screen "752_Profinet_IO_System" 1280x800, template "Top_Header"
   on GenerateScreen: SetTag("UserDiag_HmiData_actIOSystem", 1)
   on ClearScreen: SetTag("UserDiag_HmiData_actIOSystem", -2)
   TextField "Text field_1" at 7,121 size 149x32; Text 'IO Systeme / IO Systems'
   Button "Schaltfläche_64" at 950,700 size 250x80; TextOn 'Reset Übersicht / Reset overview'; TextOff 'Reset Übersicht / Reset overview'
      on Press: function_b14e0dd5("UserDiag_HmiData_ackStates", 0)
   ScreenModuleView "typeDevice_1" at 110,154 size 110x110; ScreenModuleType ""
      on Guid_{11997190-132388}: SetTag("UserDiag_HmiData_actDeviceOfScreen", 1); function_efd93a16("Pop-up_OverviewModules", 0, 0, -1, -1, 2); SetBit("UserDiag_HmiData_ioSlotDiagnosticsLoaded")
      Guid_{11997190-132400} <- "[0]"
      Guid_{11997190-132580} <- "[0]"
   ScreenModuleView "typeDevice_2" at 250,154 size 110x110; ScreenModuleType ""
      on Guid_{11997190-132388}: SetTag("UserDiag_HmiData_actDeviceOfScreen", 2); function_efd93a16("Pop-up_OverviewModules", 0, 0, -1, -1, 2); SetBit("UserDiag_HmiData_ioSlotDiagnosticsLoaded")
      Guid_{11997190-132400} <- "[1]"
      Guid_{11997190-132580} <- "[1]"
   ScreenModuleView "typeDevice_3" at 390,154 size 110x110; ScreenModuleType ""
      on Guid_{11997190-132388}: SetTag("UserDiag_HmiData_actDeviceOfScreen", 3); function_efd93a16("Pop-up_OverviewModules", 0, 0, -1, -1, 2); SetBit("UserDiag_HmiData_ioSlotDiagnosticsLoaded")
      Guid_{11997190-132400} <- "[2]"
      Guid_{11997190-132580} <- "[2]"
   ScreenModuleView "typeDevice_4" at 530,154 size 110x110; ScreenModuleType ""
      on Guid_{11997190-132388}: SetTag("UserDiag_HmiData_actDeviceOfScreen", 4); function_efd93a16("Pop-up_OverviewModules", 0, 0, -1, -1, 2); SetBit("UserDiag_HmiData_ioSlotDiagnosticsLoaded")
      Guid_{11997190-132400} <- "[3]"
      Guid_{11997190-132580} <- "[3]"
   ScreenModuleView "typeDevice_5" at 670,154 size 110x110; ScreenModuleType ""
      on Guid_{11997190-132388}: SetTag("UserDiag_HmiData_actDeviceOfScreen", 5); function_efd93a16("Pop-up_OverviewModules", 0, 0, -1, -1, 2); SetBit("UserDiag_HmiData_ioSlotDiagnosticsLoaded")
      Guid_{11997190-132400} <- "[4]"
      Guid_{11997190-132580} <- "[4]"
   ScreenModuleView "typeDevice_6" at 810,154 size 110x110; ScreenModuleType ""
      on Guid_{11997190-132388}: SetTag("UserDiag_HmiData_actDeviceOfScreen", 6); function_efd93a16("Pop-up_OverviewModules", 0, 0, -1, -1, 2); SetBit("UserDiag_HmiData_ioSlotDiagnosticsLoaded")
      Guid_{11997190-132400} <- "[5]"
      Guid_{11997190-132580} <- "[5]"
   ScreenModuleView "typeDevice_7" at 950,154 size 110x110; ScreenModuleType ""
      on Guid_{11997190-132388}: SetTag("UserDiag_HmiData_actDeviceOfScreen", 7); function_efd93a16("Pop-up_OverviewModules", 0, 0, -1, -1, 2); SetBit("UserDiag_HmiData_ioSlotDiagnosticsLoaded")
      Guid_{11997190-132400} <- "[6]"
      Guid_{11997190-132580} <- "[6]"
   ScreenModuleView "typeDevice_8" at 1090,154 size 110x110; ScreenModuleType ""
      on Guid_{11997190-132388}: SetTag("UserDiag_HmiData_actDeviceOfScreen", 8); function_efd93a16("Pop-up_OverviewModules", 0, 0, -1, -1, 2); SetBit("UserDiag_HmiData_ioSlotDiagnosticsLoaded")
      Guid_{11997190-132400} <- "[7]"
      Guid_{11997190-132580} <- "[7]"
   ScreenModuleView "typeDevice_9" at 110,294 size 110x110; ScreenModuleType ""
      on Guid_{11997190-132388}: SetTag("UserDiag_HmiData_actDeviceOfScreen", 9); function_efd93a16("Pop-up_OverviewModules", 0, 0, -1, -1, 2); SetBit("UserDiag_HmiData_ioSlotDiagnosticsLoaded")
      Guid_{11997190-132400} <- "[8]"
      Guid_{11997190-132580} <- "[8]"
   ScreenModuleView "typeDevice_10" at 250,294 size 110x110; ScreenModuleType ""
      on Guid_{11997190-132388}: SetTag("UserDiag_HmiData_actDeviceOfScreen", 10); function_efd93a16("Pop-up_OverviewModules", 0, 0, -1, -1, 2); SetBit("UserDiag_HmiData_ioSlotDiagnosticsLoaded")
      Guid_{11997190-132400} <- "[9]"
      Guid_{11997190-132580} <- "[9]"
   ScreenModuleView "typeDevice_11" at 390,294 size 110x110; ScreenModuleType ""
      on Guid_{11997190-132388}: SetTag("UserDiag_HmiData_actDeviceOfScreen", 11); function_efd93a16("Pop-up_OverviewModules", 0, 0, -1, -1, 2); SetBit("UserDiag_HmiData_ioSlotDiagnosticsLoaded")
      Guid_{11997190-132400} <- "[10]"
      Guid_{11997190-132580} <- "[10]"
   ScreenModuleView "typeDevice_12" at 530,294 size 110x110; ScreenModuleType ""
      on Guid_{11997190-132388}: SetTag("UserDiag_HmiData_actDeviceOfScreen", 12); function_efd93a16("Pop-up_OverviewModules", 0, 0, -1, -1, 2); SetBit("UserDiag_HmiData_ioSlotDiagnosticsLoaded")
      Guid_{11997190-132400} <- "[11]"
      Guid_{11997190-132580} <- "[11]"
   ScreenModuleView "typeDevice_13" at 670,294 size 110x110; ScreenModuleType ""
      on Guid_{11997190-132388}: SetTag("UserDiag_HmiData_actDeviceOfScreen", 13); function_efd93a16("Pop-up_OverviewModules", 0, 0, -1, -1, 2); SetBit("UserDiag_HmiData_ioSlotDiagnosticsLoaded")
      Guid_{11997190-132400} <- "[12]"
      Guid_{11997190-132580} <- "[12]"
   ScreenModuleView "typeDevice_14" at 810,294 size 110x110; ScreenModuleType ""
      on Guid_{11997190-132388}: SetTag("UserDiag_HmiData_actDeviceOfScreen", 14); function_efd93a16("Pop-up_OverviewModules", 0, 0, -1, -1, 2); SetBit("UserDiag_HmiData_ioSlotDiagnosticsLoaded")
      Guid_{11997190-132400} <- "[13]"
      Guid_{11997190-132580} <- "[13]"
   ScreenModuleView "typeDevice_15" at 950,292 size 110x110; ScreenModuleType ""
      on Guid_{11997190-132388}: SetTag("UserDiag_HmiData_actDeviceOfScreen", 15); function_efd93a16("Pop-up_OverviewModules", 0, 0, -1, -1, 2); SetBit("UserDiag_HmiData_ioSlotDiagnosticsLoaded")
      Guid_{11997190-132400} <- "[14]"
      Guid_{11997190-132580} <- "[14]"
   ScreenModuleView "typeDevice_16" at 1090,294 size 110x110; ScreenModuleType ""
      on Guid_{11997190-132388}: SetTag("UserDiag_HmiData_actDeviceOfScreen", 16); function_efd93a16("Pop-up_OverviewModules", 0, 0, -1, -1, 2); SetBit("UserDiag_HmiData_ioSlotDiagnosticsLoaded")
      Guid_{11997190-132400} <- "[15]"
      Guid_{11997190-132580} <- "[15]"
   ScreenModuleView "typeDevice_17" at 110,434 size 110x110; ScreenModuleType ""
      on Guid_{11997190-132388}: SetTag("UserDiag_HmiData_actDeviceOfScreen", 17); function_efd93a16("Pop-up_OverviewModules", 0, 0, -1, -1, 2); SetBit("UserDiag_HmiData_ioSlotDiagnosticsLoaded")
      Guid_{11997190-132400} <- "[16]"
      Guid_{11997190-132580} <- "[16]"
   ScreenModuleView "typeDevice_18" at 250,434 size 110x110; ScreenModuleType ""
      on Guid_{11997190-132388}: SetTag("UserDiag_HmiData_actDeviceOfScreen", 18); function_efd93a16("Pop-up_OverviewModules", 0, 0, -1, -1, 2); SetBit("UserDiag_HmiData_ioSlotDiagnosticsLoaded")
      Guid_{11997190-132400} <- "[17]"
      Guid_{11997190-132580} <- "[17]"
   ScreenModuleView "typeDevice_19" at 390,434 size 110x110; ScreenModuleType ""
      on Guid_{11997190-132388}: SetTag("UserDiag_HmiData_actDeviceOfScreen", 19); function_efd93a16("Pop-up_OverviewModules", 0, 0, -1, -1, 2); SetBit("UserDiag_HmiData_ioSlotDiagnosticsLoaded")
      Guid_{11997190-132400} <- "[18]"
      Guid_{11997190-132580} <- "[18]"
   ScreenModuleView "typeDevice_20" at 530,434 size 110x110; ScreenModuleType ""
      on Guid_{11997190-132388}: SetTag("UserDiag_HmiData_actDeviceOfScreen", 20); function_efd93a16("Pop-up_OverviewModules", 0, 0, -1, -1, 2); SetBit("UserDiag_HmiData_ioSlotDiagnosticsLoaded")
      Guid_{11997190-132400} <- "[19]"
      Guid_{11997190-132580} <- "[19]"
   ScreenModuleView "typeDevice_21" at 670,434 size 110x110; ScreenModuleType ""
      on Guid_{11997190-132388}: SetTag("UserDiag_HmiData_actDeviceOfScreen", 21); function_efd93a16("Pop-up_OverviewModules", 0, 0, -1, -1, 2); SetBit("UserDiag_HmiData_ioSlotDiagnosticsLoaded")
      Guid_{11997190-132400} <- "[20]"
      Guid_{11997190-132580} <- "[20]"
   ScreenModuleView "typeDevice_22" at 810,434 size 110x110; ScreenModuleType ""
      on Guid_{11997190-132388}: SetTag("UserDiag_HmiData_actDeviceOfScreen", 22); function_efd93a16("Pop-up_OverviewModules", 0, 0, -1, -1, 2); SetBit("UserDiag_HmiData_ioSlotDiagnosticsLoaded")
      Guid_{11997190-132400} <- "[21]"
      Guid_{11997190-132580} <- "[21]"
   ScreenModuleView "typeDevice_23" at 950,434 size 110x110; ScreenModuleType ""
      on Guid_{11997190-132388}: SetTag("UserDiag_HmiData_actDeviceOfScreen", 23); function_efd93a16("Pop-up_OverviewModules", 0, 0, -1, -1, 2); SetBit("UserDiag_HmiData_ioSlotDiagnosticsLoaded")
      Guid_{11997190-132400} <- "[22]"
      Guid_{11997190-132580} <- "[22]"
   ScreenModuleView "typeDevice_24" at 1090,434 size 110x110; ScreenModuleType ""
      on Guid_{11997190-132388}: SetTag("UserDiag_HmiData_actDeviceOfScreen", 24); function_efd93a16("Pop-up_OverviewModules", 0, 0, -1, -1, 2); SetBit("UserDiag_HmiData_ioSlotDiagnosticsLoaded")
      Guid_{11997190-132400} <- "[23]"
      Guid_{11997190-132580} <- "[23]"
   ScreenModuleView "typeDevice_25" at 110,574 size 110x110; ScreenModuleType ""
      on Guid_{11997190-132388}: SetTag("UserDiag_HmiData_actDeviceOfScreen", 25); function_efd93a16("Pop-up_OverviewModules", 0, 0, -1, -1, 2); SetBit("UserDiag_HmiData_ioSlotDiagnosticsLoaded")
      Guid_{11997190-132400} <- "[24]"
      Guid_{11997190-132580} <- "[24]"
   ScreenModuleView "typeDevice_26" at 250,574 size 110x110; ScreenModuleType ""
      on Guid_{11997190-132388}: SetTag("UserDiag_HmiData_actDeviceOfScreen", 26); function_efd93a16("Pop-up_OverviewModules", 0, 0, -1, -1, 2); SetBit("UserDiag_HmiData_ioSlotDiagnosticsLoaded")
      Guid_{11997190-132400} <- "[25]"
      Guid_{11997190-132580} <- "[25]"
   ScreenModuleView "typeDevice_27" at 390,574 size 110x110; ScreenModuleType ""
      on Guid_{11997190-132388}: SetTag("UserDiag_HmiData_actDeviceOfScreen", 27); function_efd93a16("Pop-up_OverviewModules", 0, 0, -1, -1, 2); SetBit("UserDiag_HmiData_ioSlotDiagnosticsLoaded")
      Guid_{11997190-132400} <- "[26]"
      Guid_{11997190-132580} <- "[26]"
   ScreenModuleView "typeDevice_28" at 530,574 size 110x110; ScreenModuleType ""
      on Guid_{11997190-132388}: SetTag("UserDiag_HmiData_actDeviceOfScreen", 28); function_efd93a16("Pop-up_OverviewModules", 0, 0, -1, -1, 2); SetBit("UserDiag_HmiData_ioSlotDiagnosticsLoaded")
      Guid_{11997190-132400} <- "[27]"
      Guid_{11997190-132580} <- "[27]"
   ScreenModuleView "typeDevice_29" at 670,574 size 110x110; ScreenModuleType ""
      on Guid_{11997190-132388}: SetTag("UserDiag_HmiData_actDeviceOfScreen", 29); function_efd93a16("Pop-up_OverviewModules", 0, 0, -1, -1, 2); SetBit("UserDiag_HmiData_ioSlotDiagnosticsLoaded")
      Guid_{11997190-132400} <- "[28]"
      Guid_{11997190-132580} <- "[28]"
   ScreenModuleView "typeDevice_30" at 810,574 size 110x110; ScreenModuleType ""
      on Guid_{11997190-132388}: SetTag("UserDiag_HmiData_actDeviceOfScreen", 30); function_efd93a16("Pop-up_OverviewModules", 0, 0, -1, -1, 2); SetBit("UserDiag_HmiData_ioSlotDiagnosticsLoaded")
      Guid_{11997190-132400} <- "[29]"
      Guid_{11997190-132580} <- "[29]"
   ScreenModuleView "typeDevice_31" at 950,574 size 110x110; ScreenModuleType ""
      on Guid_{11997190-132388}: SetTag("UserDiag_HmiData_actDeviceOfScreen", 31); function_efd93a16("Pop-up_OverviewModules", 0, 0, -1, -1, 2); SetBit("UserDiag_HmiData_ioSlotDiagnosticsLoaded")
      Guid_{11997190-132400} <- "[30]"
      Guid_{11997190-132580} <- "[30]"
   ScreenModuleView "typeDevice_32" at 1090,574 size 110x110; ScreenModuleType ""
      on Guid_{11997190-132388}: SetTag("UserDiag_HmiData_actDeviceOfScreen", 32); function_efd93a16("Pop-up_OverviewModules", 0, 0, -1, -1, 2); SetBit("UserDiag_HmiData_ioSlotDiagnosticsLoaded")
      Guid_{11997190-132400} <- "[31]"
      Guid_{11997190-132580} <- "[31]"
   Button "Schaltfläche_3" at 810,700 size 110x80; TextOn 'Legende / Legend'; TextOff 'Legende / Legend'
      on Click: function_efd93a16("Pop-up_Legend", 0, 0, -1, -1, 2)
   Button "Schaltfläche_4" at 110,700 size 110x80; TextOn 'Filter'; TextOff 'Filter'
      on Click: InvertBit("UserDiag_HmiData_filterErrorDevices")
      Appearance <- "UserDiag_HmiData_filterErrorDevices"
   TextField "Text field_2" at 122,160 size 86x25; Text 'Device 1'
   TextField "Text field_3" at 261,160 size 86x25; Text 'Device 2'
   TextField "Text field_4" at 401,160 size 86x25; Text 'Device 3'
   TextField "Text field_5" at 541,160 size 86x25; Text 'Device 4'
   TextField "Text field_6" at 681,160 size 86x25; Text 'Device 5'
   TextField "Text field_7" at 821,160 size 86x25; Text 'Device 6'
   TextField "Text field_8" at 961,160 size 86x25; Text 'Device 7'
   TextField "Text field_9" at 1101,160 size 86x25; Text 'Device 8'
   TextField "Text field_10" at 122,301 size 86x25; Text 'Device 9'
   TextField "Text field_11" at 256,301 size 98x25; Text 'Device 10'
   TextField "Text field_12" at 395,301 size 98x25; Text 'Device 11'
   TextField "Text field_13" at 535,301 size 98x25; Text 'Device 12'
   TextField "Text field_14" at 675,301 size 98x25; Text 'Device 13'
   TextField "Text field_15" at 815,301 size 98x25; Text 'Device 14'
   TextField "Text field_16" at 955,302 size 98x25; Text 'Device 15'
   TextField "Text field_17" at 256,301 size 98x25; Text 'Device 10'
   TextField "Text field_18" at 1096,303 size 98x25; Text 'Device 16'
   TextField "Text field_19" at 116,441 size 98x25; Text 'Device 17'
   TextField "Text field_20" at 256,442 size 98x25; Text 'Device 18'
   TextField "Text field_21" at 396,442 size 98x25; Text 'Device 19'
   TextField "Text field_22" at 536,442 size 98x25; Text 'Device 20'
   TextField "Text field_23" at 676,442 size 98x25; Text 'Device 21'
   TextField "Text field_24" at 816,442 size 98x25; Text 'Device 22'
   TextField "Text field_25" at 956,442 size 98x25; Text 'Device 23'
   TextField "Text field_26" at 1096,442 size 98x25; Text 'Device 24'
   TextField "Text field_27" at 116,583 size 98x25; Text 'Device 25'
   TextField "Text field_28" at 255,583 size 98x25; Text 'Device 26'
   TextField "Text field_29" at 395,583 size 98x25; Text 'Device 27'
   TextField "Text field_30" at 535,583 size 98x25; Text 'Device 28'
   TextField "Text field_31" at 675,583 size 98x25; Text 'Device 29'
   TextField "Text field_32" at 815,583 size 98x25; Text 'Device 30'
   TextField "Text field_33" at 955,583 size 98x25; Text 'Device 31'
   TextField "Text field_34" at 1095,583 size 98x25; Text 'Device 32'
   Button "Button_19" at 524,717 size 123x83; TextOn 'LINE_OVERVIEW_1 PROFINET DIAGNOSTIC MESSAGES'; TextOff 'LINE_OVERVIEW_1 PROFINET DIAGNOSTIC MESSAGES'
      on Click: ActivateScreen("753_Topic_003.0_Messages", 0)
   Button "Button_3" at 383,717 size 123x83; TextOn 'LINE_OVERVIEW_1 PROFINET DIAGNOSTIC MESSAGES'; TextOff 'LINE_OVERVIEW_1 PROFINET PLC DIAGNOSTIC'
      on Click: ActivateScreen("751_Topic_001.0_PLC", 0)
   Rectangle "Rectangle_2" at 20,323 size 60x97
      Appearance <- "UserDiag_HmiData_errorAtLowerScreen"
   Rectangle "Rectangle_5" at 20,420 size 60x97
      Appearance <- "UserDiag_HmiData_errorAtUpperScreen"
   IOField "I/O field_1" at 20,396 size 60x50; FormatPattern 99
      ProcessValue <- "UserDiag_HmiData_actScreenDevices"
   GraphicView "Graphic view_3" at 36,480 size 27x30; Picture "Down_Hell"
   GraphicView "Graphic view_4" at 36,328 size 27x30; Picture "Up_Hell"
   Button "Button_1" at 20,458 size 60x60; TextOff 'Text'
      on Click: "IncActScreenDev"()
   Button "Button_2" at 20,323 size 60x60; TextOff 'Text'
      on Click: "DecActScreenDev"()
   Group "Group" at 187,117 size 180x34; TextList "Text_list_IO_System"
   Rectangle "Rectangle_1" at 187,117 size 180x34
      Appearance <- "[0]"
   Rectangle "Rectangle_4" at 187,117 size 180x34
      Appearance <- "UserDiag_HmiData_actIOSystem"
   SymbolicIOField "Symbolic I/O field_2" at 187,117 size 180x34; TextOn '1'; TextOff '0'; TextList "Text_list_IO_System"
      ProcessValue <- "ioSystem1"
   Button "Schaltfläche_1" at 187,117 size 180x34; TextOff 'Text'
      on Click: SetTag("UserDiag_HmiData_actIOSystem", 1); SetTag("UserDiag_HmiData_actScreenDevices", 1)

screen "753_Topic_003.0_Messages" 1280x800, template "Top_Header"
   AlarmView "Alarm view_1" at 40,120 size 1160x574

screen "2004 - PLC Web Server Diag" 1280x800, template "Top_Header"
   on GenerateScreen: SetTag("PLC_IP_Address", 'http://172.16.0.1')
   HTMLBrowser "HTML browser_1" at 0,120 size 1280x580
      Address <- "PLC_IP_Address"
   TextField "Text field_1" at 0,720 size 168x25; Text 'PLC IP Address :'
   IOField "I/O field_1" at 148,717 size 280x32; FormatPattern ??????????????????????????????
      ProcessValue <- "PLC_IP_Address"

screen "2010 - HMI Functions" 1280x800, template "Top_Header"
   Button "Schaltfläche_1" at 645,206 size 100x100; TextOff 'Transfer'
      on Release: function_bb44b551(2)
      Appearance <- "Always_OFF_HMI"
   Button "Schaltfläche_2" at 755,324 size 100x100; TextOff 'Runtime beenden Stop Runtime'
      on Release: StopRuntime(0)
      Appearance <- "Always_OFF_HMI"
   Button "Schaltfläche_3" at 535,206 size 100x100; TextOff 'Offline'
      on Release: function_bb44b551(1)
      Appearance <- "Always_OFF_HMI"
   Button "Schaltfläche_4" at 425,206 size 100x100; TextOff 'Online'
      on Release: function_bb44b551(0)
      Appearance <- "Always_OFF_HMI"
   Button "Schaltfläche_5" at 425,324 size 100x100; TextOff 'Kalibriere Touchscreen Calibrate'
      on Release: function_bc3e350c()
      Appearance <- "Always_OFF_HMI"
   Button "Schaltfläche_8" at 645,324 size 100x100; TextOff 'Systemsteuerung Control Panel'
      on Release: function_f34a74f3()
      Appearance <- "Always_OFF_HMI"
   Button "Button_1" at 755,206 size 100x100; TextOff 'On Screen Keyboard'
      on Release: function_d6caf649(0)
      Appearance <- "Always_OFF_HMI"
   Button "Schaltfläche_6" at 535,324 size 100x100; TextOff 'Kalibriere Touchscreen Clean Screen'
      on Release: function_be740847(30)
      Appearance <- "Always_OFF_HMI"

screen "2011 - User Administration" 1280x800, template "Top_Header"
   UserView "User view_1" at 0,120 size 1280x580

screen "2003 - System Diag" 1280x800, template "Top_Header"
   SysDiagControl "System diagnostics view_1" at 0,120 size 1280x580

screen "710_ALL_CARRIER_STATUS" 1280x800, template "Top_Header"
   on GenerateScreen: "SDC_EMS_STATUS"('SDC\DB_SDC_EMS\_Intern_EMS_Nr'); "SDC_TS_REFERENCE"("SDC\DB_SDC_EMS\EMS[XXX].TS_STAT.VAL.SEK"); SetTag("SDC\DB_SDC_EMS\HMI[XX].BILD_Nr", 728); "SDC_EMS_TA_STATUS"("HMI_EMS_Nr"); SetTag("SDC\_intern_Bildnummer", 728)
   on ClearScreen: SetTag("SDC\DB_SDC_EMS\HMI[XX].BILD_Nr", 0)
   Button "Button_1" at 13,169 size 80x46; TextOff 'EMS 1'
      on Release: ActivateScreen("711_CARRIER_STATUS", 0)
      on Press: SetTag("HMI_EMS_Nr", 1)
      Appearance <- "DB16_EMS_Status_EMS_DeviceStates.DeviceStates_Condition_HMI[1]"
      ObjectEnable <- "DB16_EMS_Status_EMS_DeviceStates.DeviceStates_Condition_HMI[1]"
   Button "Button_2" at 96,169 size 80x46; TextOff 'EMS 2'
      on Release: ActivateScreen("711_CARRIER_STATUS", 0)
      on Press: SetTag("HMI_EMS_Nr", 2)
      Appearance <- "DB16_EMS_Status_EMS_DeviceStates.DeviceStates_Condition_HMI[2]"
      ObjectEnable <- "DB16_EMS_Status_EMS_DeviceStates.DeviceStates_Condition_HMI[2]"
   Button "Button_3" at 180,169 size 80x46; TextOff 'EMS 3'
      on Release: ActivateScreen("711_CARRIER_STATUS", 0)
      on Press: SetTag("HMI_EMS_Nr", 3)
      Appearance <- "DB16_EMS_Status_EMS_DeviceStates.DeviceStates_Condition_HMI[3]"
      ObjectEnable <- "DB16_EMS_Status_EMS_DeviceStates.DeviceStates_Condition_HMI[3]"
   Button "Button_4" at 263,169 size 80x46; TextOff 'EMS 4'
      on Release: ActivateScreen("711_CARRIER_STATUS", 0)
      on Press: SetTag("HMI_EMS_Nr", 4)
      Appearance <- "DB16_EMS_Status_EMS_DeviceStates.DeviceStates_Condition_HMI[4]"
      ObjectEnable <- "DB16_EMS_Status_EMS_DeviceStates.DeviceStates_Condition_HMI[4]"
   Button "Button_5" at 346,169 size 80x46; TextOff 'EMS 5'
      on Release: ActivateScreen("711_CARRIER_STATUS", 0)
      on Press: SetTag("HMI_EMS_Nr", 5)
      Appearance <- "DB16_EMS_Status_EMS_DeviceStates.DeviceStates_Condition_HMI[5]"
      ObjectEnable <- "DB16_EMS_Status_EMS_DeviceStates.DeviceStates_Condition_HMI[5]"
   Button "Button_6" at 429,169 size 80x46; TextOff 'EMS 6'
      on Release: ActivateScreen("711_CARRIER_STATUS", 0)
      on Press: SetTag("HMI_EMS_Nr", 6)
      Appearance <- "DB16_EMS_Status_EMS_DeviceStates.DeviceStates_Condition_HMI[6]"
      ObjectEnable <- "DB16_EMS_Status_EMS_DeviceStates.DeviceStates_Condition_HMI[6]"
   Button "Button_7" at 512,169 size 80x46; TextOff 'EMS 7'
      on Release: ActivateScreen("711_CARRIER_STATUS", 0)
      on Press: SetTag("HMI_EMS_Nr", 7)
      Appearance <- "DB16_EMS_Status_EMS_DeviceStates.DeviceStates_Condition_HMI[7]"
      ObjectEnable <- "DB16_EMS_Status_EMS_DeviceStates.DeviceStates_Condition_HMI[7]"
   Button "Button_8" at 595,169 size 80x46; TextOff 'EMS 8'
      on Release: ActivateScreen("711_CARRIER_STATUS", 0)
      on Press: SetTag("HMI_EMS_Nr", 8)
      Appearance <- "DB16_EMS_Status_EMS_DeviceStates.DeviceStates_Condition_HMI[8]"
      ObjectEnable <- "DB16_EMS_Status_EMS_DeviceStates.DeviceStates_Condition_HMI[8]"
   Button "Button_9" at 678,169 size 80x46; TextOff 'EMS 9'
      on Release: ActivateScreen("711_CARRIER_STATUS", 0)
      on Press: SetTag("HMI_EMS_Nr", 9)
      Appearance <- "DB16_EMS_Status_EMS_DeviceStates.DeviceStates_Condition_HMI[9]"
      ObjectEnable <- "DB16_EMS_Status_EMS_DeviceStates.DeviceStates_Condition_HMI[9]"
   Button "Button_10" at 761,169 size 80x46; TextOff 'EMS 10'
      on Release: ActivateScreen("711_CARRIER_STATUS", 0)
      on Press: SetTag("HMI_EMS_Nr", 10)
      Appearance <- "DB16_EMS_Status_EMS_DeviceStates.DeviceStates_Condition_HMI[10]"
      ObjectEnable <- "DB16_EMS_Status_EMS_DeviceStates.DeviceStates_Condition_HMI[10]"
   Button "Button_11" at 845,169 size 80x46; TextOff 'EMS 11'
      on Release: ActivateScreen("711_CARRIER_STATUS", 0)
      on Press: SetTag("HMI_EMS_Nr", 11)
      Appearance <- "DB16_EMS_Status_EMS_DeviceStates.DeviceStates_Condition_HMI[11]"
      ObjectEnable <- "DB16_EMS_Status_EMS_DeviceStates.DeviceStates_Condition_HMI[11]"
   Button "Button_12" at 928,169 size 80x46; TextOff 'EMS 12'
      on Release: ActivateScreen("711_CARRIER_STATUS", 0)
      on Press: SetTag("HMI_EMS_Nr", 12)
      Appearance <- "DB16_EMS_Status_EMS_DeviceStates.DeviceStates_Condition_HMI[12]"
      ObjectEnable <- "DB16_EMS_Status_EMS_DeviceStates.DeviceStates_Condition_HMI[12]"
   Button "Button_13" at 1011,169 size 80x46; TextOff 'EMS 13'
      on Release: ActivateScreen("711_CARRIER_STATUS", 0)
      on Press: SetTag("HMI_EMS_Nr", 13)
      Appearance <- "DB16_EMS_Status_EMS_DeviceStates.DeviceStates_Condition_HMI[13]"
      ObjectEnable <- "DB16_EMS_Status_EMS_DeviceStates.DeviceStates_Condition_HMI[13]"
   Button "Button_14" at 1094,169 size 80x46; TextOff 'EMS 14'
      on Release: ActivateScreen("711_CARRIER_STATUS", 0)
      on Press: SetTag("HMI_EMS_Nr", 14)
      Appearance <- "DB16_EMS_Status_EMS_DeviceStates.DeviceStates_Condition_HMI[14]"
      ObjectEnable <- "DB16_EMS_Status_EMS_DeviceStates.DeviceStates_Condition_HMI[14]"
   Button "Button_15" at 1178,169 size 80x46; TextOff 'EMS 15'
      on Release: ActivateScreen("711_CARRIER_STATUS", 0)
      on Press: SetTag("HMI_EMS_Nr", 15)
      Appearance <- "DB16_EMS_Status_EMS_DeviceStates.DeviceStates_Condition_HMI[15]"
      ObjectEnable <- "DB16_EMS_Status_EMS_DeviceStates.DeviceStates_Condition_HMI[15]"
   Button "Button_16" at 13,250 size 80x46; TextOff 'EMS 16'
      on Release: ActivateScreen("711_CARRIER_STATUS", 0)
      on Press: SetTag("HMI_EMS_Nr", 16)
      ObjectEnable <- "DB16_EMS_Status_EMS_DeviceStates.DeviceStates_Condition_HMI[16]"
      Appearance <- "[16]"
   Button "Button_17" at 96,250 size 80x46; TextOff 'EMS 17'
      on Release: ActivateScreen("711_CARRIER_STATUS", 0)
      on Press: SetTag("HMI_EMS_Nr", 17)
      Appearance <- "DB16_EMS_Status_EMS_DeviceStates.DeviceStates_Condition_HMI[17]"
      ObjectEnable <- "DB16_EMS_Status_EMS_DeviceStates.DeviceStates_Condition_HMI[17]"
   Button "Button_18" at 180,250 size 80x46; TextOff 'EMS 18'
      on Release: ActivateScreen("711_CARRIER_STATUS", 0)
      on Press: SetTag("HMI_EMS_Nr", 18)
      Appearance <- "DB16_EMS_Status_EMS_DeviceStates.DeviceStates_Condition_HMI[18]"
      ObjectEnable <- "DB16_EMS_Status_EMS_DeviceStates.DeviceStates_Condition_HMI[18]"
   Button "Button_19" at 263,250 size 80x46; TextOff 'EMS 19'
      on Release: ActivateScreen("711_CARRIER_STATUS", 0)
      on Press: SetTag("HMI_EMS_Nr", 19)
      Appearance <- "DB16_EMS_Status_EMS_DeviceStates.DeviceStates_Condition_HMI[19]"
      ObjectEnable <- "DB16_EMS_Status_EMS_DeviceStates.DeviceStates_Condition_HMI[19]"
   Button "Button_20" at 346,250 size 80x46; TextOff 'EMS 20'
      on Release: ActivateScreen("711_CARRIER_STATUS", 0)
      on Press: SetTag("HMI_EMS_Nr", 20)
      Appearance <- "DB16_EMS_Status_EMS_DeviceStates.DeviceStates_Condition_HMI[20]"
      ObjectEnable <- "DB16_EMS_Status_EMS_DeviceStates.DeviceStates_Condition_HMI[20]"
   Button "Button_21" at 429,250 size 80x46; TextOff 'EMS 21'
      on Release: ActivateScreen("711_CARRIER_STATUS", 0)
      on Press: SetTag("HMI_EMS_Nr", 21)
      Appearance <- "DB16_EMS_Status_EMS_DeviceStates.DeviceStates_Condition_HMI[21]"
      ObjectEnable <- "DB16_EMS_Status_EMS_DeviceStates.DeviceStates_Condition_HMI[21]"
   Button "Button_22" at 512,250 size 80x46; TextOff 'EMS 22'
      on Release: ActivateScreen("711_CARRIER_STATUS", 0)
      on Press: SetTag("HMI_EMS_Nr", 22)
      Appearance <- "DB16_EMS_Status_EMS_DeviceStates.DeviceStates_Condition_HMI[22]"
      ObjectEnable <- "DB16_EMS_Status_EMS_DeviceStates.DeviceStates_Condition_HMI[22]"
   Button "Button_23" at 595,250 size 80x46; TextOff 'EMS 23'
      on Release: ActivateScreen("711_CARRIER_STATUS", 0)
      on Press: SetTag("HMI_EMS_Nr", 23)
      Appearance <- "DB16_EMS_Status_EMS_DeviceStates.DeviceStates_Condition_HMI[23]"
      ObjectEnable <- "DB16_EMS_Status_EMS_DeviceStates.DeviceStates_Condition_HMI[23]"
   Button "Button_24" at 678,250 size 80x46; TextOff 'EMS 24'
      on Release: ActivateScreen("711_CARRIER_STATUS", 0)
      on Press: SetTag("HMI_EMS_Nr", 24)
      Appearance <- "DB16_EMS_Status_EMS_DeviceStates.DeviceStates_Condition_HMI[24]"
      ObjectEnable <- "DB16_EMS_Status_EMS_DeviceStates.DeviceStates_Condition_HMI[24]"
   Button "Button_25" at 761,250 size 80x46; TextOff 'EMS 25'
      on Release: ActivateScreen("711_CARRIER_STATUS", 0)
      on Press: SetTag("HMI_EMS_Nr", 25)
      Appearance <- "DB16_EMS_Status_EMS_DeviceStates.DeviceStates_Condition_HMI[25]"
      ObjectEnable <- "DB16_EMS_Status_EMS_DeviceStates.DeviceStates_Condition_HMI[25]"
   Button "Button_26" at 845,250 size 80x46; TextOff 'EMS 26'
      on Release: ActivateScreen("711_CARRIER_STATUS", 0)
      on Press: SetTag("HMI_EMS_Nr", 26)
      Appearance <- "DB16_EMS_Status_EMS_DeviceStates.DeviceStates_Condition_HMI[26]"
      ObjectEnable <- "DB16_EMS_Status_EMS_DeviceStates.DeviceStates_Condition_HMI[26]"
   Button "Button_27" at 928,250 size 80x46; TextOff 'EMS 27'
      on Release: ActivateScreen("711_CARRIER_STATUS", 0)
      on Press: SetTag("HMI_EMS_Nr", 27)
      Appearance <- "DB16_EMS_Status_EMS_DeviceStates.DeviceStates_Condition_HMI[27]"
      ObjectEnable <- "DB16_EMS_Status_EMS_DeviceStates.DeviceStates_Condition_HMI[27]"
   Button "Button_28" at 1011,250 size 80x46; TextOff 'EMS 28'
      on Release: ActivateScreen("711_CARRIER_STATUS", 0)
      on Press: SetTag("HMI_EMS_Nr", 28)
      Appearance <- "DB16_EMS_Status_EMS_DeviceStates.DeviceStates_Condition_HMI[28]"
      ObjectEnable <- "DB16_EMS_Status_EMS_DeviceStates.DeviceStates_Condition_HMI[28]"
   Button "Button_29" at 1094,250 size 80x46; TextOff 'EMS 29'
      on Release: ActivateScreen("711_CARRIER_STATUS", 0)
      on Press: SetTag("HMI_EMS_Nr", 29)
      Appearance <- "DB16_EMS_Status_EMS_DeviceStates.DeviceStates_Condition_HMI[29]"
      ObjectEnable <- "DB16_EMS_Status_EMS_DeviceStates.DeviceStates_Condition_HMI[29]"
   Button "Button_30" at 1178,250 size 80x46; TextOff 'EMS 30'
      on Release: ActivateScreen("711_CARRIER_STATUS", 0)
      on Press: SetTag("HMI_EMS_Nr", 30)
      Appearance <- "DB16_EMS_Status_EMS_DeviceStates.DeviceStates_Condition_HMI[30]"
      ObjectEnable <- "DB16_EMS_Status_EMS_DeviceStates.DeviceStates_Condition_HMI[30]"
   Button "Button_31" at 13,331 size 80x46; TextOff 'EMS 31'
      on Release: ActivateScreen("711_CARRIER_STATUS", 0)
      on Press: SetTag("HMI_EMS_Nr", 31)
      ObjectEnable <- "DB16_EMS_Status_EMS_DeviceStates.DeviceStates_Condition_HMI[31]"
      Appearance <- "[31]"
   Button "Button_32" at 96,331 size 80x46; TextOff 'EMS 32'
      on Release: ActivateScreen("711_CARRIER_STATUS", 0)
      on Press: SetTag("HMI_EMS_Nr", 32)
      ObjectEnable <- "DB16_EMS_Status_EMS_DeviceStates.DeviceStates_Condition_HMI[32]"
      Appearance <- "[32]"
   Button "Button_33" at 180,331 size 80x46; TextOff 'EMS 33'
      on Release: ActivateScreen("711_CARRIER_STATUS", 0)
      on Press: SetTag("HMI_EMS_Nr", 33)
      ObjectEnable <- "DB16_EMS_Status_EMS_DeviceStates.DeviceStates_Condition_HMI[33]"
      Appearance <- "[33]"
   Button "Button_34" at 263,331 size 80x46; TextOff 'EMS 34'
      on Release: ActivateScreen("711_CARRIER_STATUS", 0)
      on Press: SetTag("HMI_EMS_Nr", 34)
      ObjectEnable <- "DB16_EMS_Status_EMS_DeviceStates.DeviceStates_Condition_HMI[34]"
      Appearance <- "[34]"
   Button "Button_35" at 346,331 size 80x46; TextOff 'EMS 35'
      on Release: ActivateScreen("711_CARRIER_STATUS", 0)
      on Press: SetTag("HMI_EMS_Nr", 35)
      ObjectEnable <- "DB16_EMS_Status_EMS_DeviceStates.DeviceStates_Condition_HMI[35]"
      Appearance <- "[35]"
   Button "Button_36" at 429,331 size 80x46; TextOff 'EMS 36'
      on Release: ActivateScreen("711_CARRIER_STATUS", 0)
      on Press: SetTag("HMI_EMS_Nr", 36)
      ObjectEnable <- "DB16_EMS_Status_EMS_DeviceStates.DeviceStates_Condition_HMI[36]"
      Appearance <- "[36]"
   Button "Button_37" at 512,331 size 80x46; TextOff 'EMS 37'
      on Release: ActivateScreen("711_CARRIER_STATUS", 0)
      on Press: SetTag("HMI_EMS_Nr", 37)
      ObjectEnable <- "DB16_EMS_Status_EMS_DeviceStates.DeviceStates_Condition_HMI[37]"
      Appearance <- "[37]"
   Button "Button_38" at 595,331 size 80x46; TextOff 'EMS 38'
      on Release: ActivateScreen("711_CARRIER_STATUS", 0)
      on Press: SetTag("HMI_EMS_Nr", 38)
      ObjectEnable <- "DB16_EMS_Status_EMS_DeviceStates.DeviceStates_Condition_HMI[38]"
      Appearance <- "[38]"
   Button "Button_39" at 678,331 size 80x46; TextOff 'EMS 39'
      on Release: ActivateScreen("711_CARRIER_STATUS", 0)
      on Press: SetTag("HMI_EMS_Nr", 39)
      ObjectEnable <- "DB16_EMS_Status_EMS_DeviceStates.DeviceStates_Condition_HMI[39]"
      Appearance <- "[39]"
   Button "Button_40" at 761,331 size 80x46; TextOff 'EMS 40'
      on Release: ActivateScreen("711_CARRIER_STATUS", 0)
      on Press: SetTag("HMI_EMS_Nr", 40)
      ObjectEnable <- "DB16_EMS_Status_EMS_DeviceStates.DeviceStates_Condition_HMI[40]"
      Appearance <- "[40]"
   Button "Button_41" at 845,331 size 80x46; TextOff 'EMS 41'
      on Release: ActivateScreen("711_CARRIER_STATUS", 0)
      on Press: SetTag("HMI_EMS_Nr", 41)
      ObjectEnable <- "DB16_EMS_Status_EMS_DeviceStates.DeviceStates_Condition_HMI[41]"
      Appearance <- "[41]"
   Button "Button_42" at 928,331 size 80x46; TextOff 'EMS 42'
      on Release: ActivateScreen("711_CARRIER_STATUS", 0)
      on Press: SetTag("HMI_EMS_Nr", 42)
      ObjectEnable <- "DB16_EMS_Status_EMS_DeviceStates.DeviceStates_Condition_HMI[42]"
      Appearance <- "[42]"
   Button "Button_43" at 1011,331 size 80x46; TextOff 'EMS 43'
      on Release: ActivateScreen("711_CARRIER_STATUS", 0)
      on Press: SetTag("HMI_EMS_Nr", 43)
      ObjectEnable <- "DB16_EMS_Status_EMS_DeviceStates.DeviceStates_Condition_HMI[43]"
      Appearance <- "[43]"
   Button "Button_44" at 1094,331 size 80x46; TextOff 'EMS 44'
      on Release: ActivateScreen("711_CARRIER_STATUS", 0)
      on Press: SetTag("HMI_EMS_Nr", 44)
      ObjectEnable <- "DB16_EMS_Status_EMS_DeviceStates.DeviceStates_Condition_HMI[44]"
      Appearance <- "[44]"
   Button "Button_45" at 1178,331 size 80x46; TextOff 'EMS 45'
      on Release: ActivateScreen("711_CARRIER_STATUS", 0)
      on Press: SetTag("HMI_EMS_Nr", 45)
      ObjectEnable <- "DB16_EMS_Status_EMS_DeviceStates.DeviceStates_Condition_HMI[45]"
      Appearance <- "[45]"
   Button "Button_46" at 13,412 size 80x46; TextOff 'EMS 46'
      on Release: ActivateScreen("711_CARRIER_STATUS", 0)
      on Press: SetTag("HMI_EMS_Nr", 46)
      ObjectEnable <- "DB16_EMS_Status_EMS_DeviceStates.DeviceStates_Condition_HMI[46]"
      Appearance <- "[46]"
   Button "Button_47" at 96,412 size 80x46; TextOff 'EMS 47'
      on Release: ActivateScreen("711_CARRIER_STATUS", 0)
      on Press: SetTag("HMI_EMS_Nr", 47)
      ObjectEnable <- "DB16_EMS_Status_EMS_DeviceStates.DeviceStates_Condition_HMI[47]"
      Appearance <- "[47]"
   Button "Button_48" at 180,412 size 80x46; TextOff 'EMS 48'
      on Release: ActivateScreen("711_CARRIER_STATUS", 0)
      on Press: SetTag("HMI_EMS_Nr", 48)
      ObjectEnable <- "DB16_EMS_Status_EMS_DeviceStates.DeviceStates_Condition_HMI[48]"
      Appearance <- "[48]"
   Button "Button_49" at 263,412 size 80x46; TextOff 'EMS 49'
      on Release: ActivateScreen("711_CARRIER_STATUS", 0)
      on Press: SetTag("HMI_EMS_Nr", 49)
      ObjectEnable <- "DB16_EMS_Status_EMS_DeviceStates.DeviceStates_Condition_HMI[49]"
      Appearance <- "[49]"
   Button "Button_50" at 346,412 size 80x46; TextOff 'EMS 50'
      on Release: ActivateScreen("711_CARRIER_STATUS", 0)
      on Press: SetTag("HMI_EMS_Nr", 50)
      ObjectEnable <- "DB16_EMS_Status_EMS_DeviceStates.DeviceStates_Condition_HMI[50]"
      Appearance <- "[50]"
   Button "Button_51" at 429,412 size 80x46; TextOff 'EMS 51'
      on Release: ActivateScreen("711_CARRIER_STATUS", 0)
      on Press: SetTag("HMI_EMS_Nr", 51)
      ObjectEnable <- "DB16_EMS_Status_EMS_DeviceStates.DeviceStates_Condition_HMI[51]"
      Appearance <- "[51]"
   Button "Button_52" at 512,412 size 80x46; TextOff 'EMS 52'
      on Release: ActivateScreen("711_CARRIER_STATUS", 0)
      on Press: SetTag("HMI_EMS_Nr", 52)
      ObjectEnable <- "DB16_EMS_Status_EMS_DeviceStates.DeviceStates_Condition_HMI[52]"
      Appearance <- "[52]"
   Button "Button_53" at 595,412 size 80x46; TextOff 'EMS 53'
      on Release: ActivateScreen("711_CARRIER_STATUS", 0)
      on Press: SetTag("HMI_EMS_Nr", 53)
      ObjectEnable <- "DB16_EMS_Status_EMS_DeviceStates.DeviceStates_Condition_HMI[53]"
      Appearance <- "[53]"
   Button "Button_54" at 678,412 size 80x46; TextOff 'EMS 54'
      on Release: ActivateScreen("711_CARRIER_STATUS", 0)
      on Press: SetTag("HMI_EMS_Nr", 54)
      ObjectEnable <- "DB16_EMS_Status_EMS_DeviceStates.DeviceStates_Condition_HMI[54]"
      Appearance <- "[54]"
   Button "Button_55" at 761,412 size 80x46; TextOff 'EMS 55'
      on Release: ActivateScreen("711_CARRIER_STATUS", 0)
      on Press: SetTag("HMI_EMS_Nr", 55)
      ObjectEnable <- "DB16_EMS_Status_EMS_DeviceStates.DeviceStates_Condition_HMI[55]"
      Appearance <- "[55]"
   Button "Button_56" at 845,412 size 80x46; TextOff 'EMS 56'
      on Release: ActivateScreen("711_CARRIER_STATUS", 0)
      on Press: SetTag("HMI_EMS_Nr", 56)
      ObjectEnable <- "DB16_EMS_Status_EMS_DeviceStates.DeviceStates_Condition_HMI[56]"
      Appearance <- "[56]"
   Button "Button_57" at 928,412 size 80x46; TextOff 'EMS 57'
      on Release: ActivateScreen("711_CARRIER_STATUS", 0)
      on Press: SetTag("HMI_EMS_Nr", 57)
      ObjectEnable <- "DB16_EMS_Status_EMS_DeviceStates.DeviceStates_Condition_HMI[57]"
      Appearance <- "[57]"
   Button "Button_58" at 1011,412 size 80x46; TextOff 'EMS 58'
      on Release: ActivateScreen("711_CARRIER_STATUS", 0)
      on Press: SetTag("HMI_EMS_Nr", 58)
      ObjectEnable <- "DB16_EMS_Status_EMS_DeviceStates.DeviceStates_Condition_HMI[58]"
      Appearance <- "[58]"
   Button "Button_59" at 1094,412 size 80x46; TextOff 'EMS 59'
      on Release: ActivateScreen("711_CARRIER_STATUS", 0)
      on Press: SetTag("HMI_EMS_Nr", 59)
      ObjectEnable <- "DB16_EMS_Status_EMS_DeviceStates.DeviceStates_Condition_HMI[59]"
      Appearance <- "[59]"
   Button "Button_60" at 1178,412 size 80x46; TextOff 'EMS 60'
      on Release: ActivateScreen("711_CARRIER_STATUS", 0)
      on Press: SetTag("HMI_EMS_Nr", 60)
      ObjectEnable <- "DB16_EMS_Status_EMS_DeviceStates.DeviceStates_Condition_HMI[60]"
      Appearance <- "[60]"
   Button "Button_61" at 13,493 size 80x46; TextOff 'EMS 61'
      on Release: ActivateScreen("711_CARRIER_STATUS", 0)
      on Press: SetTag("HMI_EMS_Nr", 61)
      ObjectEnable <- "DB16_EMS_Status_EMS_DeviceStates.DeviceStates_Condition_HMI[61]"
      Appearance <- "[61]"
   Button "Button_62" at 96,493 size 80x46; TextOff 'EMS 62'
      on Release: ActivateScreen("711_CARRIER_STATUS", 0)
      on Press: SetTag("HMI_EMS_Nr", 62)
      ObjectEnable <- "DB16_EMS_Status_EMS_DeviceStates.DeviceStates_Condition_HMI[62]"
      Appearance <- "[62]"
   Button "Button_63" at 180,493 size 80x46; TextOff 'EMS 63'
      on Release: ActivateScreen("711_CARRIER_STATUS", 0)
      on Press: SetTag("HMI_EMS_Nr", 63)
      ObjectEnable <- "DB16_EMS_Status_EMS_DeviceStates.DeviceStates_Condition_HMI[63]"
      Appearance <- "[63]"
   Button "Button_64" at 263,493 size 80x46; TextOff 'EMS 64'
      on Release: ActivateScreen("711_CARRIER_STATUS", 0)
      on Press: SetTag("HMI_EMS_Nr", 64)
      ObjectEnable <- "DB16_EMS_Status_EMS_DeviceStates.DeviceStates_Condition_HMI[64]"
      Appearance <- "[64]"
   Button "Button_65" at 346,493 size 80x46; TextOff 'EMS 65'
      on Release: ActivateScreen("711_CARRIER_STATUS", 0)
      on Press: SetTag("HMI_EMS_Nr", 65)
      ObjectEnable <- "DB16_EMS_Status_EMS_DeviceStates.DeviceStates_Condition_HMI[65]"
      Appearance <- "[65]"
   Button "Button_66" at 429,493 size 80x46; TextOff 'EMS 66'
      on Release: ActivateScreen("711_CARRIER_STATUS", 0)
      on Press: SetTag("HMI_EMS_Nr", 66)
      ObjectEnable <- "DB16_EMS_Status_EMS_DeviceStates.DeviceStates_Condition_HMI[66]"
      Appearance <- "[66]"
   Button "Button_67" at 512,493 size 80x46; TextOff 'EMS 67'
      on Release: ActivateScreen("711_CARRIER_STATUS", 0)
      on Press: SetTag("HMI_EMS_Nr", 67)
      ObjectEnable <- "DB16_EMS_Status_EMS_DeviceStates.DeviceStates_Condition_HMI[67]"
      Appearance <- "[67]"
   Button "Button_68" at 595,493 size 80x46; TextOff 'EMS 68'
      on Release: ActivateScreen("711_CARRIER_STATUS", 0)
      on Press: SetTag("HMI_EMS_Nr", 68)
      ObjectEnable <- "DB16_EMS_Status_EMS_DeviceStates.DeviceStates_Condition_HMI[68]"
      Appearance <- "[68]"
   Button "Button_69" at 678,493 size 80x46; TextOff 'EMS 69'
      on Release: ActivateScreen("711_CARRIER_STATUS", 0)
      on Press: SetTag("HMI_EMS_Nr", 69)
      ObjectEnable <- "DB16_EMS_Status_EMS_DeviceStates.DeviceStates_Condition_HMI[69]"
      Appearance <- "[69]"
   Button "Button_70" at 761,493 size 80x46; TextOff 'EMS 70'
      on Release: ActivateScreen("711_CARRIER_STATUS", 0)
      on Press: SetTag("HMI_EMS_Nr", 70)
      ObjectEnable <- "DB16_EMS_Status_EMS_DeviceStates.DeviceStates_Condition_HMI[70]"
      Appearance <- "[70]"
   Button "Button_71" at 845,493 size 80x46; TextOff 'EMS 71'
      on Release: ActivateScreen("711_CARRIER_STATUS", 0)
      on Press: SetTag("HMI_EMS_Nr", 71)
      ObjectEnable <- "DB16_EMS_Status_EMS_DeviceStates.DeviceStates_Condition_HMI[71]"
      Appearance <- "[71]"
   Button "Button_72" at 928,493 size 80x46; TextOff 'EMS 72'
      on Release: ActivateScreen("711_CARRIER_STATUS", 0)
      on Press: SetTag("HMI_EMS_Nr", 72)
      ObjectEnable <- "DB16_EMS_Status_EMS_DeviceStates.DeviceStates_Condition_HMI[72]"
      Appearance <- "[72]"
   Button "Button_73" at 1011,493 size 80x46; TextOff 'EMS 73'
      on Release: ActivateScreen("711_CARRIER_STATUS", 0)
      on Press: SetTag("HMI_EMS_Nr", 73)
      ObjectEnable <- "DB16_EMS_Status_EMS_DeviceStates.DeviceStates_Condition_HMI[73]"
      Appearance <- "[73]"
   Button "Button_74" at 1094,493 size 80x46; TextOff 'EMS 74'
      on Release: ActivateScreen("711_CARRIER_STATUS", 0)
      on Press: SetTag("HMI_EMS_Nr", 74)
      ObjectEnable <- "DB16_EMS_Status_EMS_DeviceStates.DeviceStates_Condition_HMI[74]"
      Appearance <- "[74]"
   Button "Button_75" at 1178,493 size 80x46; TextOff 'EMS 75'
      on Release: ActivateScreen("711_CARRIER_STATUS", 0)
      on Press: SetTag("HMI_EMS_Nr", 75)
      ObjectEnable <- "DB16_EMS_Status_EMS_DeviceStates.DeviceStates_Condition_HMI[75]"
      Appearance <- "[75]"
   Button "Button_76" at 13,574 size 80x46; TextOff 'EMS 76'
      on Release: ActivateScreen("711_CARRIER_STATUS", 0)
      on Press: SetTag("HMI_EMS_Nr", 76)
      ObjectEnable <- "DB16_EMS_Status_EMS_DeviceStates.DeviceStates_Condition_HMI[76]"
      Appearance <- "[76]"
   Button "Button_77" at 96,574 size 80x46; TextOff 'EMS 77'
      on Release: ActivateScreen("711_CARRIER_STATUS", 0)
      on Press: SetTag("HMI_EMS_Nr", 77)
      ObjectEnable <- "DB16_EMS_Status_EMS_DeviceStates.DeviceStates_Condition_HMI[77]"
      Appearance <- "[77]"
   Button "Button_78" at 180,574 size 80x46; TextOff 'EMS 78'
      on Release: ActivateScreen("711_CARRIER_STATUS", 0)
      on Press: SetTag("HMI_EMS_Nr", 78)
      ObjectEnable <- "DB16_EMS_Status_EMS_DeviceStates.DeviceStates_Condition_HMI[78]"